(* Logix 5000 project; controller PLC_MCC1201_220AP1 vendor 1 type 14 code 164 rev 35.11; software revision 35.00; part 18 of 25 *)
(* tags used below, declared in another part *)
   B152 : DINT[50];
   B153 : DINT[20];
   B154 : DINT[20];
   B3 : DINT[102];
   C1_ACTIVE_LAMP : ALIAS FOR N54[260].0;
   C1_NTH_IN_LMP : ALIAS FOR N54[260].10;
   C1_NTH_IN_PE : ALIAS FOR N54[260].6;
   C1_NTH_IN_SS : ALIAS FOR N54[260].2;
   C1_NTH_OUT_LMP : ALIAS FOR N54[260].9;
   C1_NTH_OUT_PE : ALIAS FOR N54[260].5;
   C1_NTH_OUT_SS : ALIAS FOR N54[260].1;
   C1_STH_IN_LMP : ALIAS FOR N54[260].12;
   C1_STH_IN_PE : ALIAS FOR N54[260].8;
   C1_STH_IN_SS : ALIAS FOR N54[260].4;
   C1_STH_OUT_LMP : ALIAS FOR N54[260].11;
   C1_STH_OUT_PE : ALIAS FOR N54[260].7;
   C1_STH_OUT_SS : ALIAS FOR N54[260].3;
   C2_ACTIVE_LAMP : ALIAS FOR N54[261].0;
   C2_NTH_IN_LMP : ALIAS FOR N54[261].10;
   C2_NTH_IN_PE : ALIAS FOR N54[261].6;
   C2_NTH_IN_SS : ALIAS FOR N54[261].2;
   C2_NTH_OUT_LMP : ALIAS FOR N54[261].9;
   C2_NTH_OUT_PE : ALIAS FOR N54[261].5;
   C2_NTH_OUT_SS : ALIAS FOR N54[261].1;
   C2_STH_IN_LMP : ALIAS FOR N54[261].12;
   C2_STH_IN_PE : ALIAS FOR N54[261].8;
   C2_STH_IN_SS : ALIAS FOR N54[261].4;
   C2_STH_OUT_LMP : ALIAS FOR N54[261].11;
   C2_STH_OUT_PE : ALIAS FOR N54[261].7;
   C2_STH_OUT_SS : ALIAS FOR N54[261].3;
   C3_ACTIVE_LAMP : ALIAS FOR N54[262].0;
   C3_NTH_IN_LMP : ALIAS FOR N54[262].10;
   C3_NTH_IN_PE : ALIAS FOR N54[262].6;
   C3_NTH_IN_SS : ALIAS FOR N54[262].2;
   C3_NTH_OUT_LMP : ALIAS FOR N54[262].9;
   C3_NTH_OUT_PE : ALIAS FOR N54[262].5;
   C3_NTH_OUT_SS : ALIAS FOR N54[262].1;
   C3_STH_IN_LMP : ALIAS FOR N54[262].12;
   C3_STH_IN_PE : ALIAS FOR N54[262].8;
   C3_STH_IN_SS : ALIAS FOR N54[262].4;
   C3_STH_OUT_LMP : ALIAS FOR N54[262].11;
   C3_STH_OUT_PE : ALIAS FOR N54[262].7;
   C3_STH_OUT_SS : ALIAS FOR N54[262].3;
   C3_STP : ALIAS FOR O[35].10;
   C5 : COUNTER[100];
   C5_ACTIVE_LAMP : ALIAS FOR N54[264].0;
   C5_NTH_IN_SS : ALIAS FOR N54[264].2;
   C5_NTH_OUT_SS : ALIAS FOR N54[264].1;
   C5_STH_IN_SS : ALIAS FOR N54[264].4;
   C5_STH_OUT_SS : ALIAS FOR N54[264].3;
   CAWSV_ON_BIT_TO_WPLC : ALIAS FOR N251[900].0;
   I : INT[128];
   MADSEN_2IN_PULS : ALIAS FOR I[12].15;
   N163 : DINT[5];
   N53 : DINT[10];
   N54 : DINT[501];
   O : INT[128];
   REL_2IN_PULSE : ALIAS FOR N54[301].1;
   REL_DATA_REQ : ALIAS FOR N54[301].0;
   RELDR_ESTOP : ALIAS FOR I[80].0;
   S : INT[128];
   Status : INT;   // INT tag to retrieve Status value through GSV created during conversion
   T160 : TIMER[100];
   T4 : TIMER[100];
   T51 : TIMER[13];
   T57 : TIMER[100];
   TONY : ALIAS FOR B3[10].15;
   WASH_AK1_CON : ALIAS FOR N54[203].4;
   WASH_AK1_CR : ALIAS FOR N54[207].4;
   WASH_AK1_RET : ALIAS FOR N54[203].3;
   WASH_AK1_SV : ALIAS FOR O[36].2;
   WASH_AK1LO_CVG : ALIAS FOR N54[206].4;
   WASH_AK1UP_CVG : ALIAS FOR N54[205].4;
   WASH_AK2_CON : ALIAS FOR N54[203].6;
   WASH_AK2_CR : ALIAS FOR N54[207].5;
   WASH_AK2_RET : ALIAS FOR N54[203].5;
   WASH_AK2_SV : ALIAS FOR O[36].0;
   WASH_AK2LO_CVG : ALIAS FOR N54[206].5;
   WASH_AK2UP_CVG : ALIAS FOR N54[205].5;
   WASH_ARK_AUTO : ALIAS FOR N54[203].1;
   WASH_ARK_MANUAL : ALIAS FOR N54[203].2;
   WASH_CR_ACK : ALIAS FOR N54[207].0;
   WASH_SPY_AUTO : ALIAS FOR N54[204].1;
   WASH_SPY_MANLMP : ALIAS FOR N54[204].9;
   WASH_SPY_MANUAL : ALIAS FOR N54[204].2;
   WASH_SPY_OFF : ALIAS FOR N54[204].4;
   WASH_SPY_ON : ALIAS FOR N54[204].3;
   WATER2_ON : ALIAS FOR O[47].8;
   WATER3_CR : ALIAS FOR N54[207].6;
   WATER3_ON : ALIAS FOR O[47].9;
(* MainProgram, continued *)

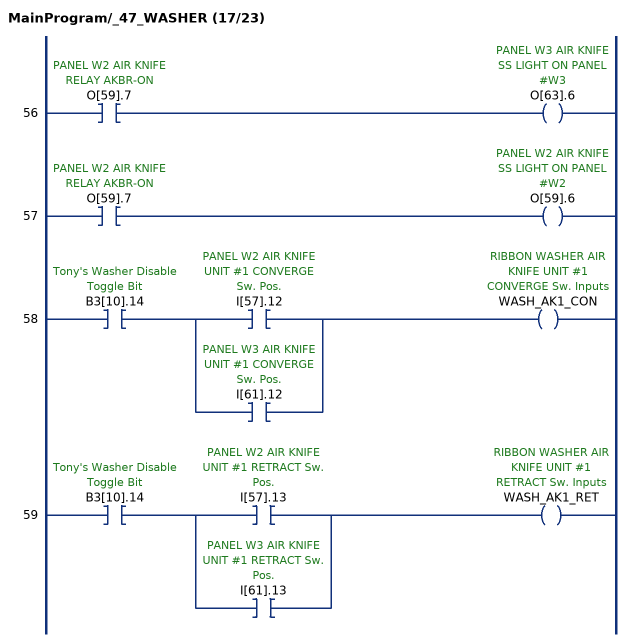
   [picture p282: MainProgram/_47_WASHER rungs 56-59]
   56: XIC(O[59].7)OTE(O[63].6);
   57: XIC(O[59].7)OTE(O[59].6);
   58: XIC(B3[10].14)[XIC(I[57].12) ,XIC(I[61].12) ]OTE(WASH_AK1_CON);
   59: XIC(B3[10].14)[XIC(I[57].13) ,XIC(I[61].13) ]OTE(WASH_AK1_RET);
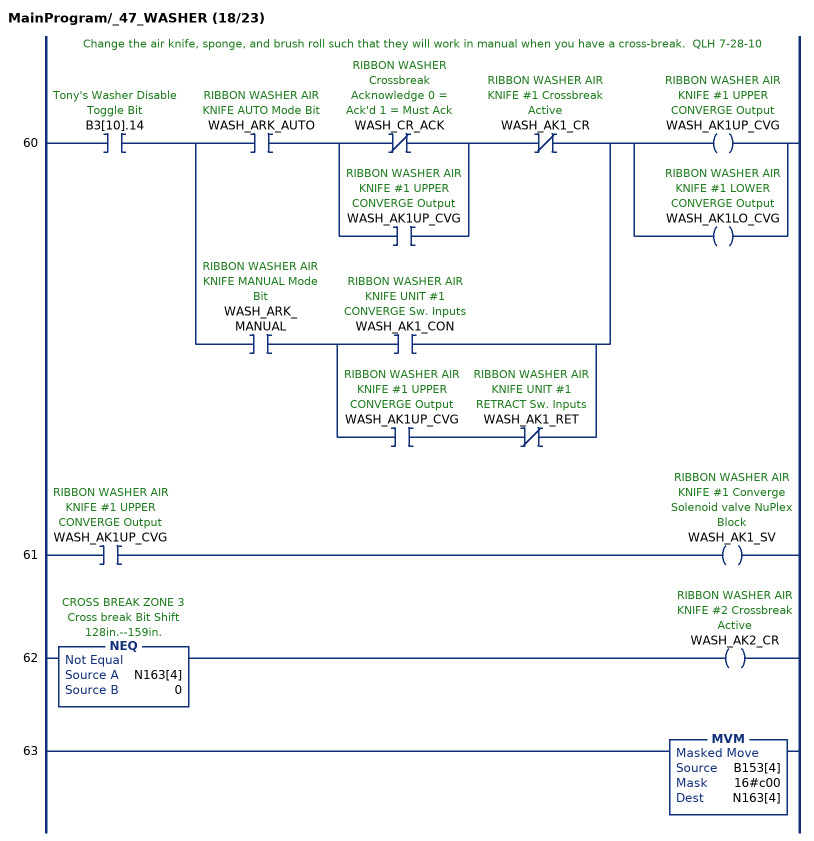
   // Change the air knife, sponge, and brush roll such that they will work in manual when you have a cross-break.  QLH 7-28-10
   60: XIC(B3[10].14)[XIC(WASH_ARK_AUTO) [XIO(WASH_CR_ACK) ,XIC(WASH_AK1UP_CVG) ] XIO(WASH_AK1_CR) ,XIC(WASH_ARK_MANUAL) [XIC(WASH_AK1_CON) ,XIC(WASH_AK1UP_CVG) XIO(WASH_AK1_RET) ] ][OTE(WASH_AK1UP_CVG) ,OTE(WASH_AK1LO_CVG) ];
   61: XIC(WASH_AK1UP_CVG)OTE(WASH_AK1_SV);
   62: NEQ(N163[4],0)OTE(WASH_AK2_CR);
   63: MVM(B153[4],16#c00,N163[4]);
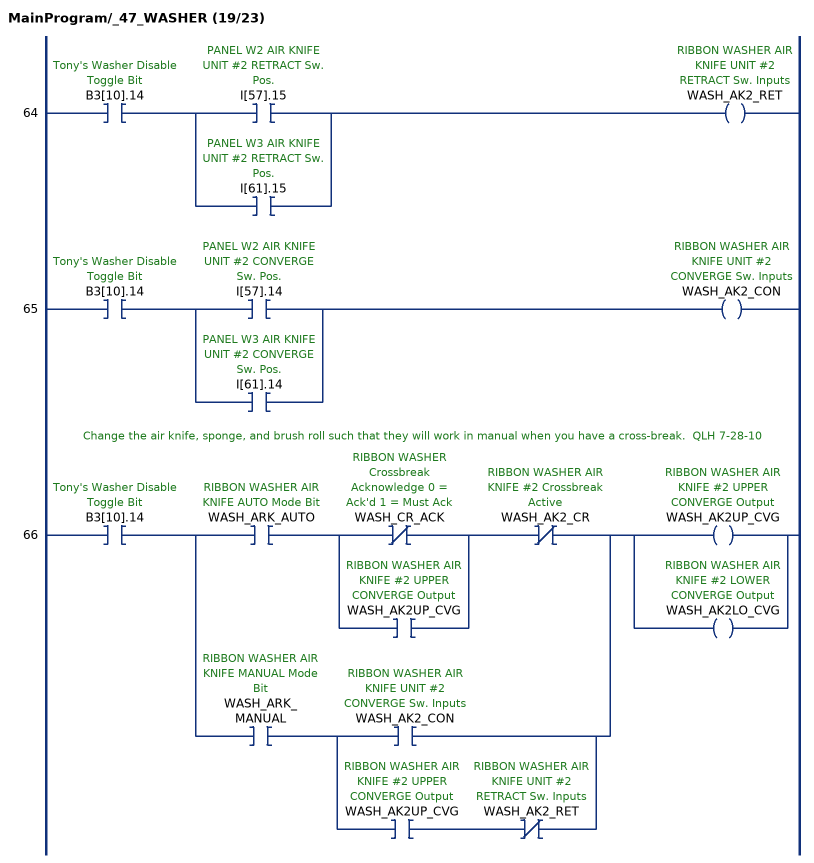
   64: XIC(B3[10].14)[XIC(I[57].15) ,XIC(I[61].15) ]OTE(WASH_AK2_RET);
   65: XIC(B3[10].14)[XIC(I[57].14) ,XIC(I[61].14) ]OTE(WASH_AK2_CON);
   // Change the air knife, sponge, and brush roll such that they will work in manual when you have a cross-break.  QLH 7-28-10
   66: XIC(B3[10].14)[XIC(WASH_ARK_AUTO) [XIO(WASH_CR_ACK) ,XIC(WASH_AK2UP_CVG) ] XIO(WASH_AK2_CR) ,XIC(WASH_ARK_MANUAL) [XIC(WASH_AK2_CON) ,XIC(WASH_AK2UP_CVG) XIO(WASH_AK2_RET) ] ][OTE(WASH_AK2UP_CVG) ,OTE(WASH_AK2LO_CVG) ];
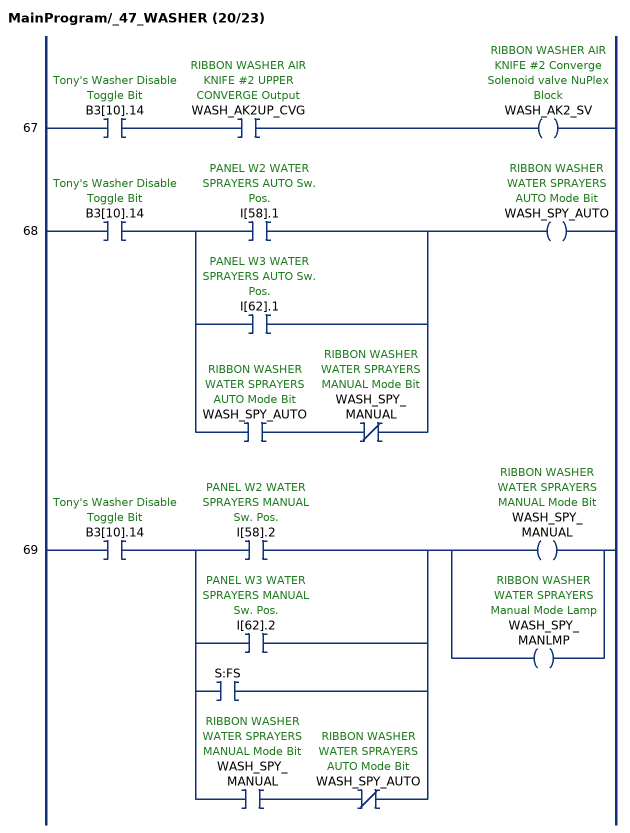
   67: XIC(B3[10].14)XIC(WASH_AK2UP_CVG)OTE(WASH_AK2_SV);
   68: XIC(B3[10].14)[[XIC(I[58].1) ,XIC(I[62].1) ] ,XIC(WASH_SPY_AUTO) XIO(WASH_SPY_MANUAL) ]OTE(WASH_SPY_AUTO);
   69: XIC(B3[10].14)[[XIC(I[58].2) ,XIC(I[62].2) ,XIC(S:FS) ] ,XIC(WASH_SPY_MANUAL) XIO(WASH_SPY_AUTO) ][OTE(WASH_SPY_MANUAL) ,OTE(WASH_SPY_MANLMP) ];
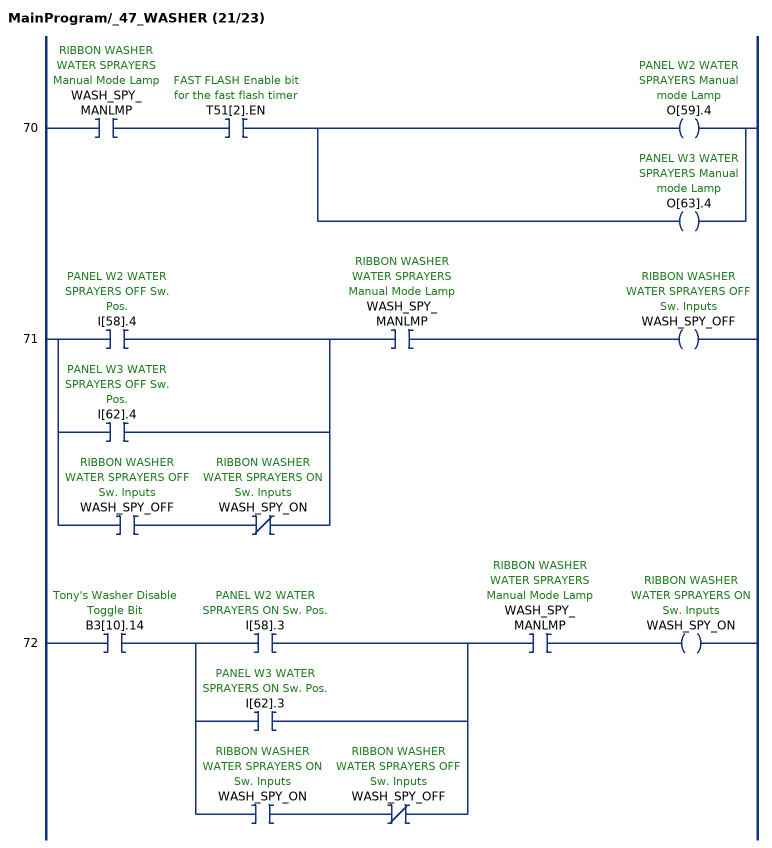
   70: XIC(WASH_SPY_MANLMP)XIC(T51[2].EN)[OTE(O[59].4) ,OTE(O[63].4) ];
   71: [[XIC(I[58].4) ,XIC(I[62].4) ] ,XIC(WASH_SPY_OFF) XIO(WASH_SPY_ON) ]XIC(WASH_SPY_MANLMP)OTE(WASH_SPY_OFF);
   72: XIC(B3[10].14)[[XIC(I[58].3) ,XIC(I[62].3) ] ,XIC(WASH_SPY_ON) XIO(WASH_SPY_OFF) ]XIC(WASH_SPY_MANLMP)OTE(WASH_SPY_ON);
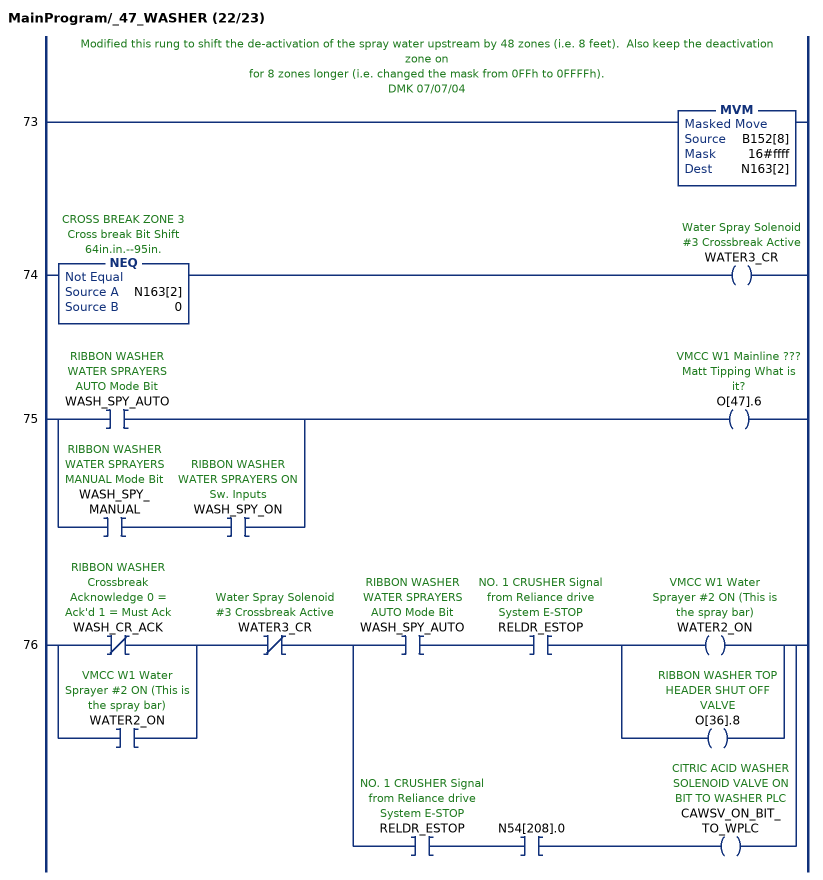
   // Modified this rung to shift the de-activation of the spray water upstream by 48 zones (i.e. 8 feet).  Also keep the deactivation zone on
   // for 8 zones longer (i.e. changed the mask from 0FFh to 0FFFFh).
   // DMK 07/07/04
   73: MVM(B152[8],16#ffff,N163[2]);
   74: NEQ(N163[2],0)OTE(WATER3_CR);
   75: [XIC(WASH_SPY_AUTO) ,XIC(WASH_SPY_MANUAL) XIC(WASH_SPY_ON) ]OTE(O[47].6);
   76: [XIO(WASH_CR_ACK) ,XIC(WATER2_ON) ]XIO(WATER3_CR)[XIC(WASH_SPY_AUTO) XIC(RELDR_ESTOP) [OTE(WATER2_ON) ,OTE(O[36].8) ] ,XIC(RELDR_ESTOP) XIC(N54[208].0) OTE(CAWSV_ON_BIT_TO_WPLC) ];
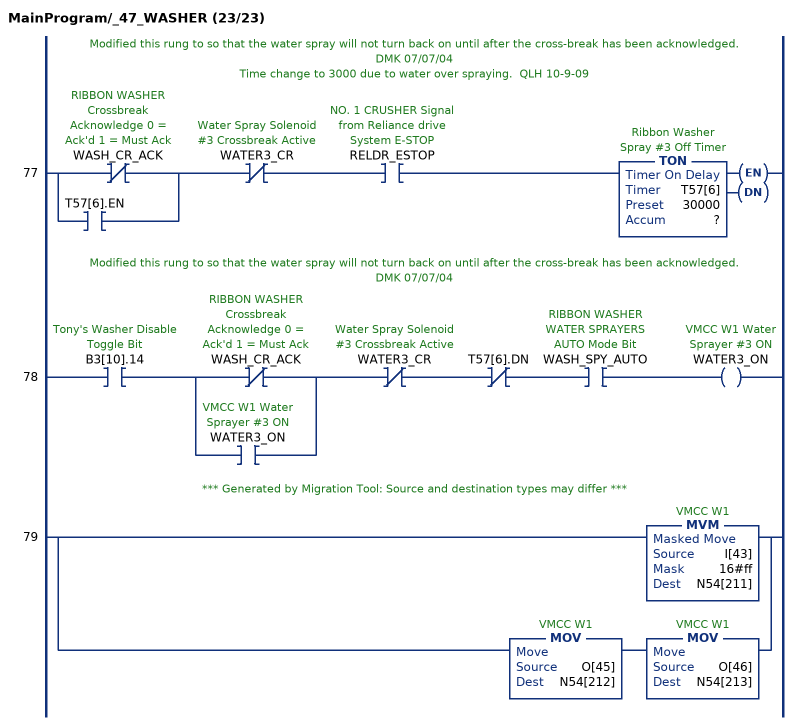
   // Modified this rung to so that the water spray will not turn back on until after the cross-break has been acknowledged.
   // DMK 07/07/04
   // Time change to 3000 due to water over spraying.  QLH 10-9-09
   77: [XIO(WASH_CR_ACK) ,XIC(T57[6].EN) ]XIO(WATER3_CR)XIC(RELDR_ESTOP)TON(T57[6],?,?);
   // Modified this rung to so that the water spray will not turn back on until after the cross-break has been acknowledged.
   // DMK 07/07/04
   78: XIC(B3[10].14)[XIO(WASH_CR_ACK) ,XIC(WATER3_ON) ]XIO(WATER3_CR)XIO(T57[6].DN)XIC(WASH_SPY_AUTO)OTE(WATER3_ON);
   // *** Generated by Migration Tool: Source and destination types may differ ***
   79: [MVM(I[43],16#ff,N54[211]) ,MOV(O[45],N54[212]) MOV(O[46],N54[213]) ];
END_ROUTINE

ROUTINE _48_IMAGE   (* ladder *)
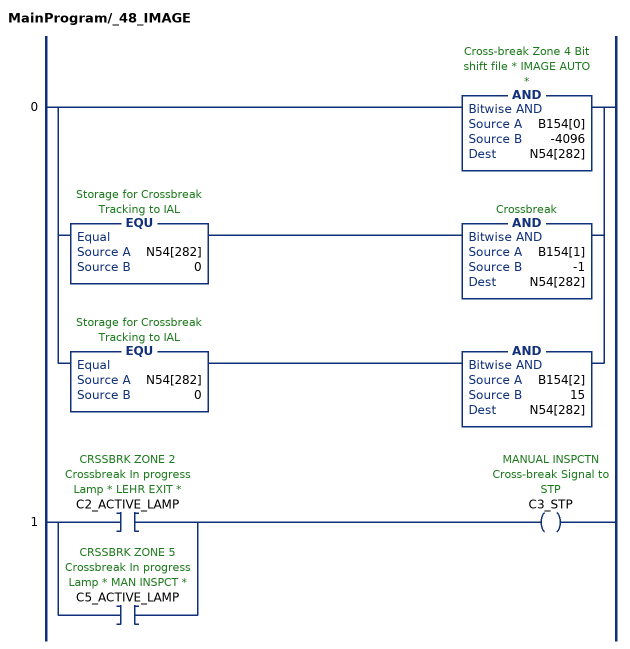
   0: [AND(B154[0],-4096,N54[282]) ,EQU(N54[282],0) AND(B154[1],-1,N54[282]) ,EQU(N54[282],0) AND(B154[2],15,N54[282]) ];
   1: [XIC(C2_ACTIVE_LAMP) ,XIC(C5_ACTIVE_LAMP) ]OTE(C3_STP);
END_ROUTINE

ROUTINE _49_INSP_REL   (* ladder *)
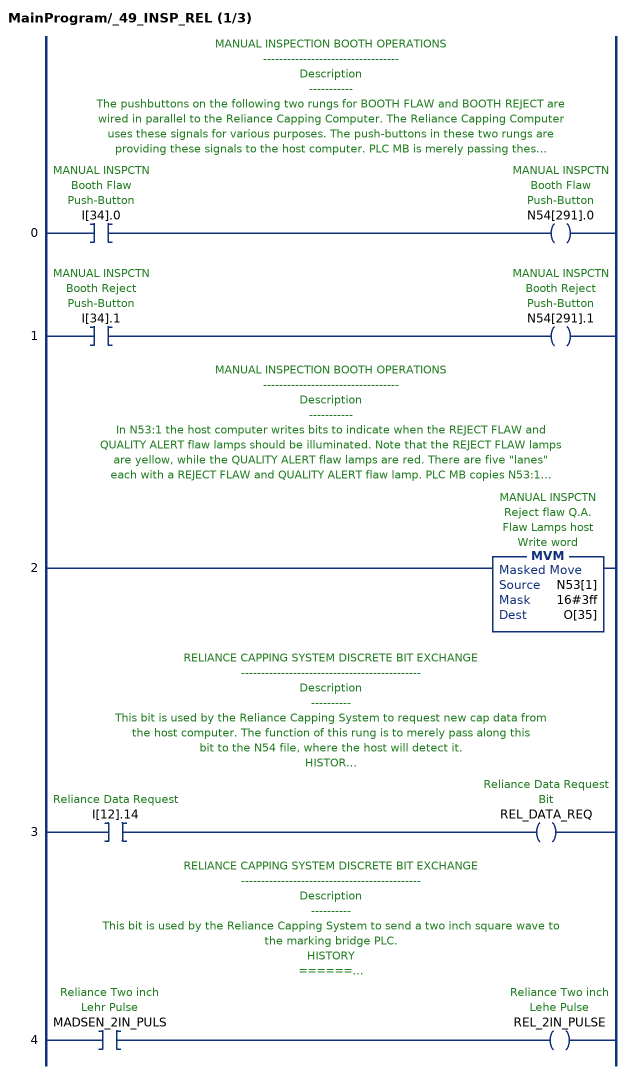
   // MANUAL INSPECTION BOOTH OPERATIONS
   // ----------------------------------
   // Description
   // -----------
   // The pushbuttons on the following two rungs for BOOTH FLAW and BOOTH REJECT are
   // wired in parallel to the Reliance Capping Computer. The Reliance Capping Computer
   // uses these signals for various purposes. The push-buttons in these two rungs are
   // providing these signals to the host computer. PLC MB is merely passing these
   // signals along to the host computer.
   // HISTORY
   // =======
   // Date       Description                                                Programmer
   // ----       -----------                                                ----------
   // 3/11/96    Added this rung and comments.                                WAS
   0: XIC(I[34].0)OTE(N54[291].0);
   1: XIC(I[34].1)OTE(N54[291].1);
   // MANUAL INSPECTION BOOTH OPERATIONS
   // ----------------------------------
   // Description
   // -----------
   // In N53:1 the host computer writes bits to indicate when the REJECT FLAW and
   // QUALITY ALERT flaw lamps should be illuminated. Note that the REJECT FLAW lamps
   // are yellow, while the QUALITY ALERT flaw lamps are red. There are five "lanes"
   // each with a REJECT FLAW and QUALITY ALERT flaw lamp. PLC MB copies N53:1,
   // the host write area, to O:043, the actual output word for the lamps.
   // HISTORY
   // =======
   // Date       Description                                                Programmer
   // ----       -----------                                                ----------
   // 3/11/96    Added this rung and comments.                                WAS
   2: MVM(N53[1],16#3ff,O[35]);
   // RELIANCE CAPPING SYSTEM DISCRETE BIT EXCHANGE
   // ---------------------------------------------
   // Description
   // ----------
   // This bit is used by the Reliance Capping System to request new cap data from
   // the host computer. The function of this rung is to merely pass along this
   // bit to the N54 file, where the host will detect it.
   // HISTORY
   // =======
   // Date       Description                                                Programmer
   // ----       -----------                                                ----------
   // 3/11/96    Discussed issue with Steve Sutter. Elected to locate This    WAS
   //            bit in local rack in case timing becomes critical.
   // 3/11/96    Added this rung and comments.                                WAS
   3: XIC(I[12].14)OTE(REL_DATA_REQ);
   // RELIANCE CAPPING SYSTEM DISCRETE BIT EXCHANGE
   // ---------------------------------------------
   // Description
   // ----------
   // This bit is used by the Reliance Capping System to send a two inch square wave to
   // the marking bridge PLC.
   // HISTORY
   // =======
   // Date       Description                                                Programmer
   // ----       -----------                                                ----------
   // 3/11/96    Discussed issue with Steve Sutter. Elected to locate This    WAS
   //            bit in local rack in case timing becomes critical.
   // 3/11/96    Added this rung and comments.                                WAS
   4: XIC(MADSEN_2IN_PULS)OTE(REL_2IN_PULSE);
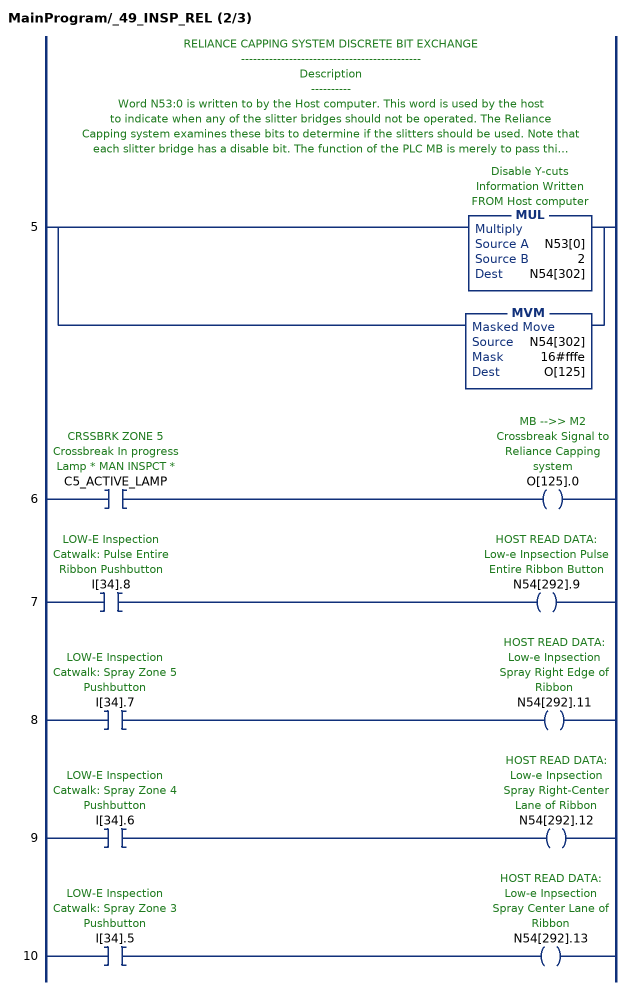
   // RELIANCE CAPPING SYSTEM DISCRETE BIT EXCHANGE
   // ---------------------------------------------
   // Description
   // ----------
   // Word N53:0 is written to by the Host computer. This word is used by the host
   // to indicate when any of the slitter bridges should not be operated. The Reliance
   // Capping system examines these bits to determine if the slitters should be used. Note that
   // each slitter bridge has a disable bit. The function of the PLC MB is merely to pass this
   // data along from the Host computer to the Reliance Capping System.
   // HISTORY
   // =======
   // Date       Description                                                Programmer
   // ----       -----------                                                ----------
   // 3/11/96    Added this rung and comments.                                WAS
   5: [MUL(N53[0],2,N54[302]) ,MVM(N54[302],16#fffe,O[125]) ];
   6: XIC(C5_ACTIVE_LAMP)OTE(O[125].0);
   7: XIC(I[34].8)OTE(N54[292].9);
   8: XIC(I[34].7)OTE(N54[292].11);
   9: XIC(I[34].6)OTE(N54[292].12);
   10: XIC(I[34].5)OTE(N54[292].13);
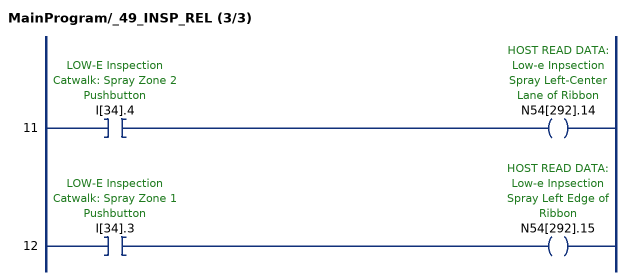
   11: XIC(I[34].4)OTE(N54[292].14);
   12: XIC(I[34].3)OTE(N54[292].15);
END_ROUTINE

ROUTINE _50_I_O_REMAP   (* ladder *)
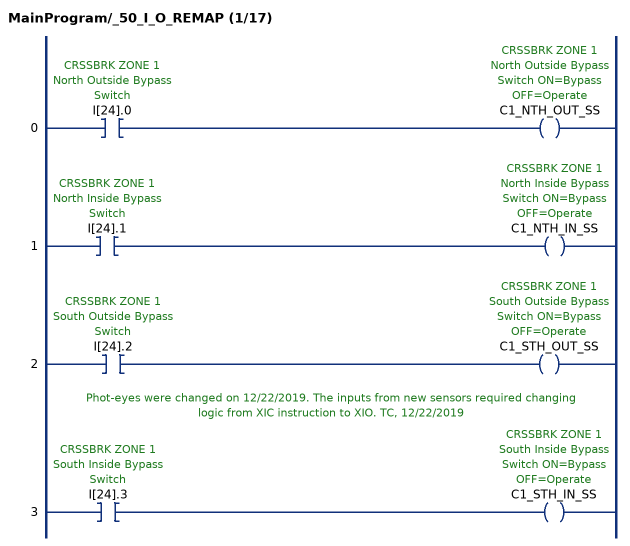
   0: XIC(I[24].0)OTE(C1_NTH_OUT_SS);
   1: XIC(I[24].1)OTE(C1_NTH_IN_SS);
   2: XIC(I[24].2)OTE(C1_STH_OUT_SS);
   // Phot-eyes were changed on 12/22/2019. The inputs from new sensors required changing logic from XIC instruction to XIO. TC, 12/22/2019
   3: XIC(I[24].3)OTE(C1_STH_IN_SS);
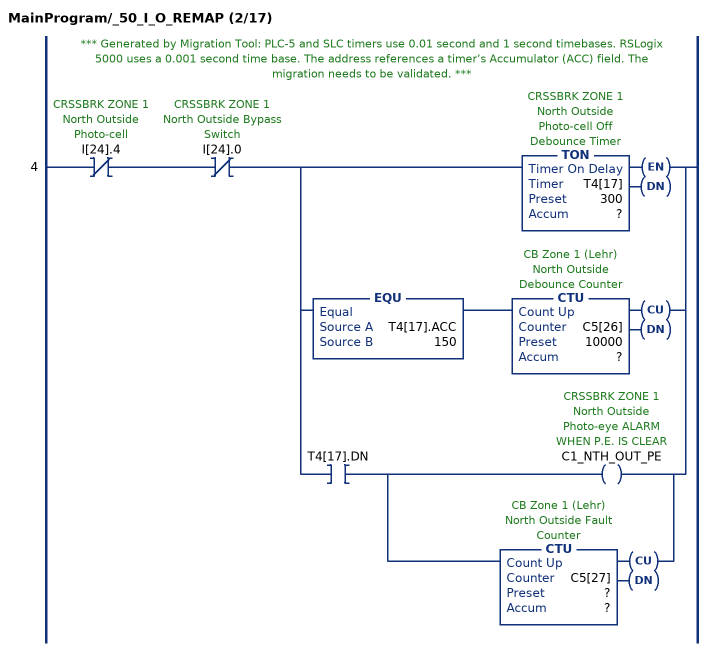
   // *** Generated by Migration Tool: PLC-5 and SLC timers use 0.01 second and 1 second timebases. RSLogix 5000 uses a 0.001 second time base. The address references a timer’s Accumulator (ACC) field. The migration needs to be validated. ***
   4: XIO(I[24].4)XIO(I[24].0)[TON(T4[17],?,?) ,EQU(T4[17].ACC,150) CTU(C5[26],?,?) ,XIC(T4[17].DN) [OTE(C1_NTH_OUT_PE) ,CTU(C5[27],?,?) ] ];
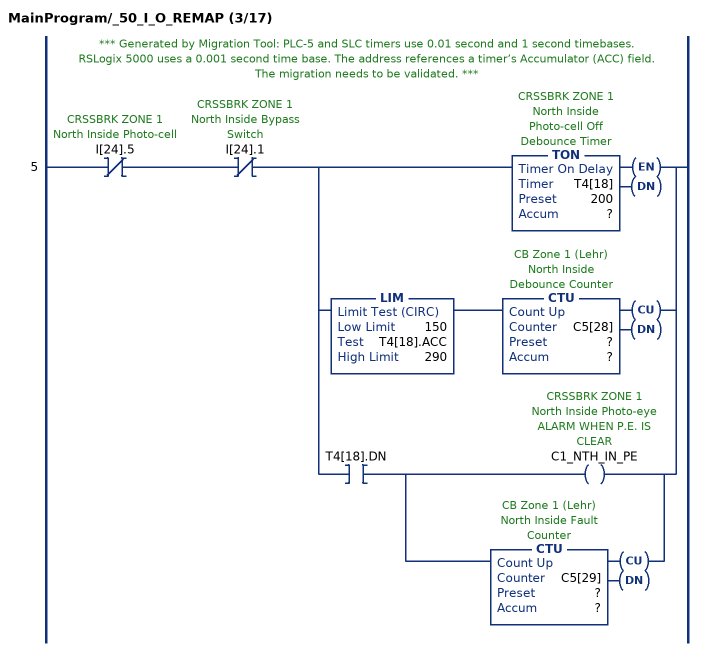
   // *** Generated by Migration Tool: PLC-5 and SLC timers use 0.01 second and 1 second timebases. RSLogix 5000 uses a 0.001 second time base. The address references a timer’s Accumulator (ACC) field. The migration needs to be validated. ***
   5: XIO(I[24].5)XIO(I[24].1)[TON(T4[18],?,?) ,LIM(150,T4[18].ACC,290) CTU(C5[28],?,?) ,XIC(T4[18].DN) [OTE(C1_NTH_IN_PE) ,CTU(C5[29],?,?) ] ];
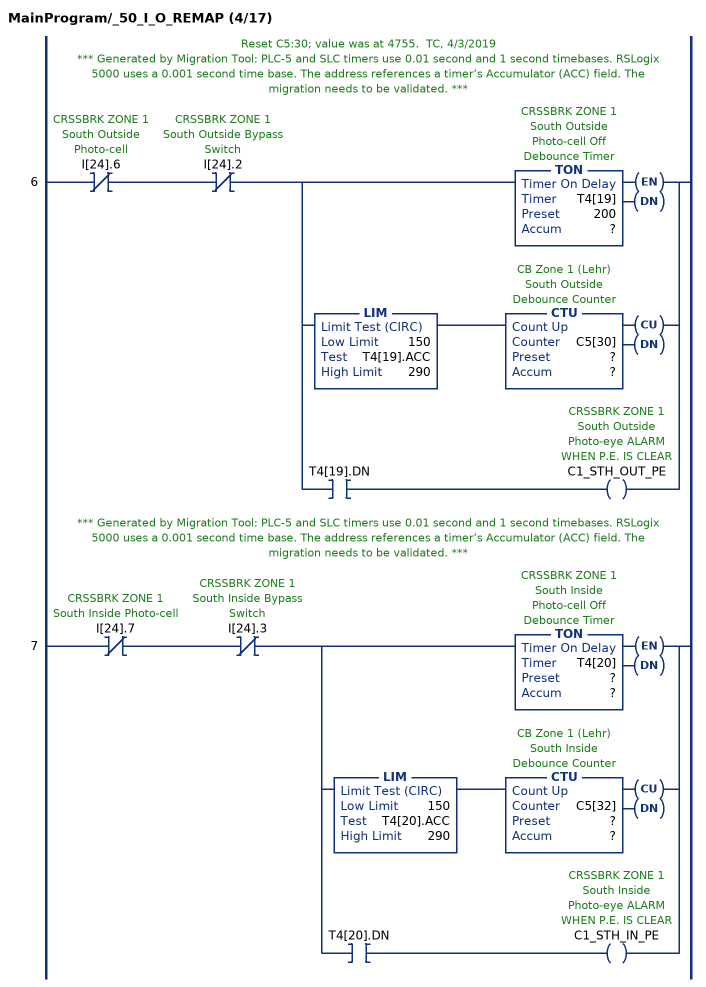
   // Reset C5:30; value was at 4755.  TC, 4/3/2019
   // *** Generated by Migration Tool: PLC-5 and SLC timers use 0.01 second and 1 second timebases. RSLogix 5000 uses a 0.001 second time base. The address references a timer’s Accumulator (ACC) field. The migration needs to be validated. ***
   6: XIO(I[24].6)XIO(I[24].2)[TON(T4[19],?,?) ,LIM(150,T4[19].ACC,290) CTU(C5[30],?,?) ,XIC(T4[19].DN) OTE(C1_STH_OUT_PE) ];
   // *** Generated by Migration Tool: PLC-5 and SLC timers use 0.01 second and 1 second timebases. RSLogix 5000 uses a 0.001 second time base. The address references a timer’s Accumulator (ACC) field. The migration needs to be validated. ***
   7: XIO(I[24].7)XIO(I[24].3)[TON(T4[20],?,?) ,LIM(150,T4[20].ACC,290) CTU(C5[32],?,?) ,XIC(T4[20].DN) OTE(C1_STH_IN_PE) ];
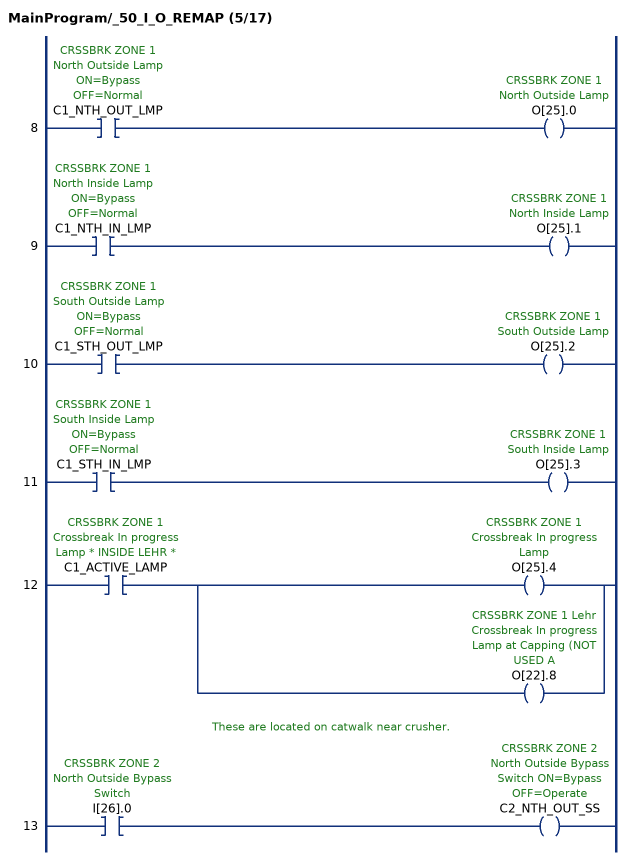
   8: XIC(C1_NTH_OUT_LMP)OTE(O[25].0);
   9: XIC(C1_NTH_IN_LMP)OTE(O[25].1);
   10: XIC(C1_STH_OUT_LMP)OTE(O[25].2);
   11: XIC(C1_STH_IN_LMP)OTE(O[25].3);
   12: XIC(C1_ACTIVE_LAMP)[OTE(O[25].4) ,OTE(O[22].8) ];
   // These are located on catwalk near crusher.
   13: XIC(I[26].0)OTE(C2_NTH_OUT_SS);
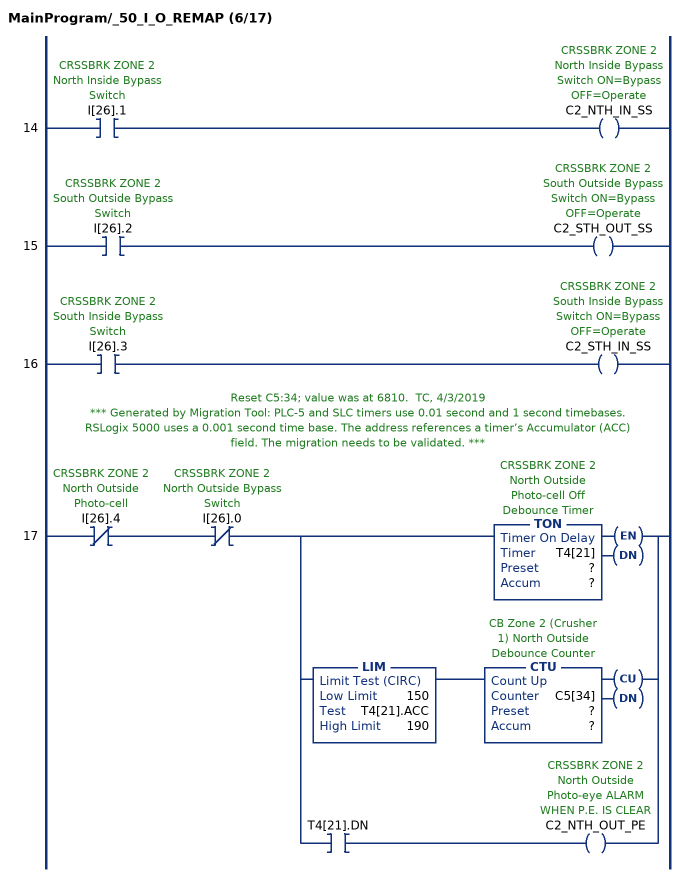
   14: XIC(I[26].1)OTE(C2_NTH_IN_SS);
   15: XIC(I[26].2)OTE(C2_STH_OUT_SS);
   16: XIC(I[26].3)OTE(C2_STH_IN_SS);
   // Reset C5:34; value was at 6810.  TC, 4/3/2019
   // *** Generated by Migration Tool: PLC-5 and SLC timers use 0.01 second and 1 second timebases. RSLogix 5000 uses a 0.001 second time base. The address references a timer’s Accumulator (ACC) field. The migration needs to be validated. ***
   17: XIO(I[26].4)XIO(I[26].0)[TON(T4[21],?,?) ,LIM(150,T4[21].ACC,190) CTU(C5[34],?,?) ,XIC(T4[21].DN) OTE(C2_NTH_OUT_PE) ];
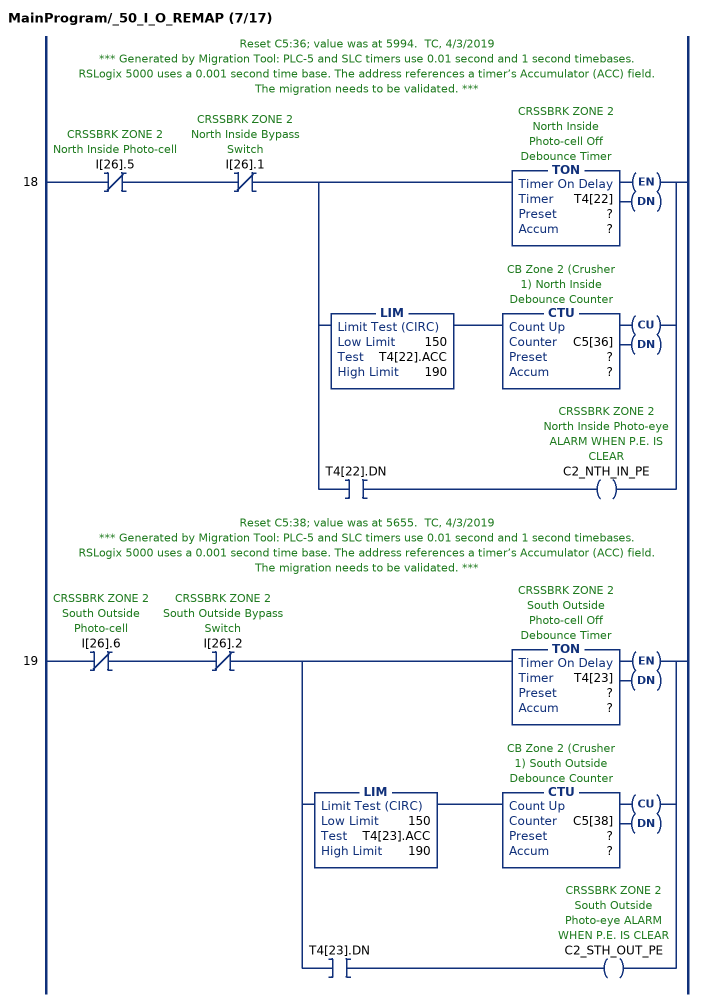
   // Reset C5:36; value was at 5994.  TC, 4/3/2019
   // *** Generated by Migration Tool: PLC-5 and SLC timers use 0.01 second and 1 second timebases. RSLogix 5000 uses a 0.001 second time base. The address references a timer’s Accumulator (ACC) field. The migration needs to be validated. ***
   18: XIO(I[26].5)XIO(I[26].1)[TON(T4[22],?,?) ,LIM(150,T4[22].ACC,190) CTU(C5[36],?,?) ,XIC(T4[22].DN) OTE(C2_NTH_IN_PE) ];
   // Reset C5:38; value was at 5655.  TC, 4/3/2019
   // *** Generated by Migration Tool: PLC-5 and SLC timers use 0.01 second and 1 second timebases. RSLogix 5000 uses a 0.001 second time base. The address references a timer’s Accumulator (ACC) field. The migration needs to be validated. ***
   19: XIO(I[26].6)XIO(I[26].2)[TON(T4[23],?,?) ,LIM(150,T4[23].ACC,190) CTU(C5[38],?,?) ,XIC(T4[23].DN) OTE(C2_STH_OUT_PE) ];
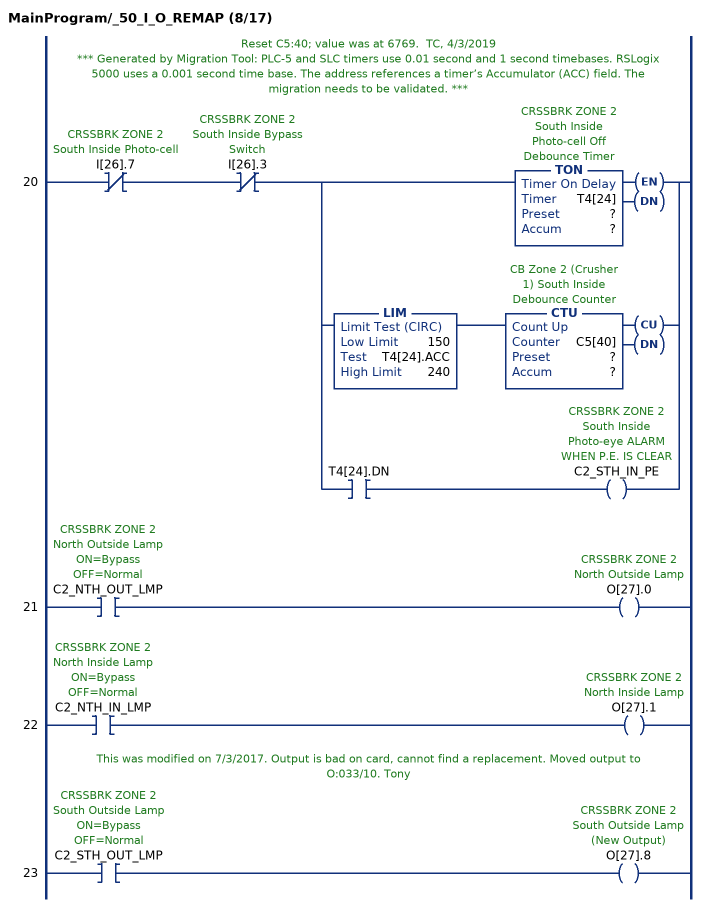
   // Reset C5:40; value was at 6769.  TC, 4/3/2019
   // *** Generated by Migration Tool: PLC-5 and SLC timers use 0.01 second and 1 second timebases. RSLogix 5000 uses a 0.001 second time base. The address references a timer’s Accumulator (ACC) field. The migration needs to be validated. ***
   20: XIO(I[26].7)XIO(I[26].3)[TON(T4[24],?,?) ,LIM(150,T4[24].ACC,240) CTU(C5[40],?,?) ,XIC(T4[24].DN) OTE(C2_STH_IN_PE) ];
   21: XIC(C2_NTH_OUT_LMP)OTE(O[27].0);
   22: XIC(C2_NTH_IN_LMP)OTE(O[27].1);
   // This was modified on 7/3/2017. Output is bad on card, cannot find a replacement. Moved output to O:033/10. Tony
   23: XIC(C2_STH_OUT_LMP)OTE(O[27].8);
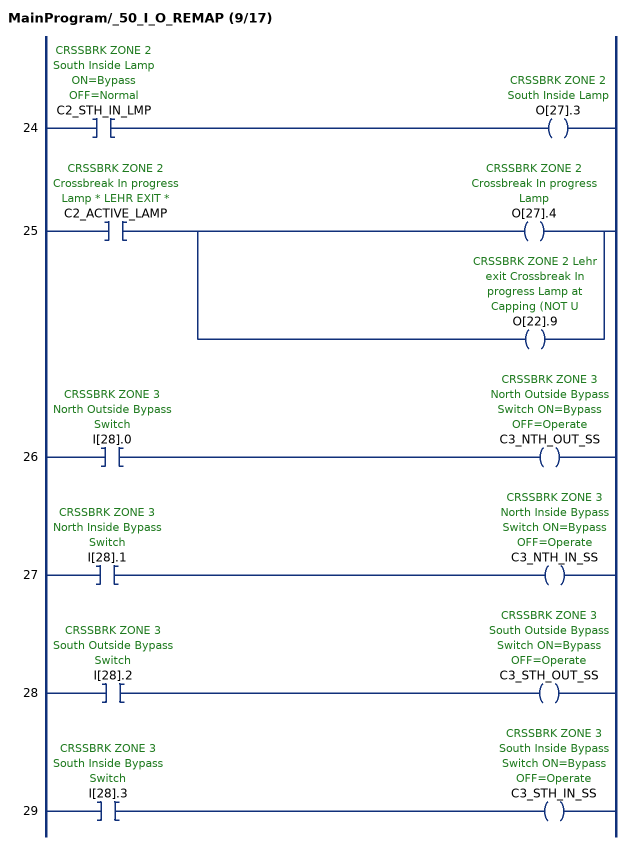
   24: XIC(C2_STH_IN_LMP)OTE(O[27].3);
   25: XIC(C2_ACTIVE_LAMP)[OTE(O[27].4) ,OTE(O[22].9) ];
   26: XIC(I[28].0)OTE(C3_NTH_OUT_SS);
   27: XIC(I[28].1)OTE(C3_NTH_IN_SS);
   28: XIC(I[28].2)OTE(C3_STH_OUT_SS);
   29: XIC(I[28].3)OTE(C3_STH_IN_SS);
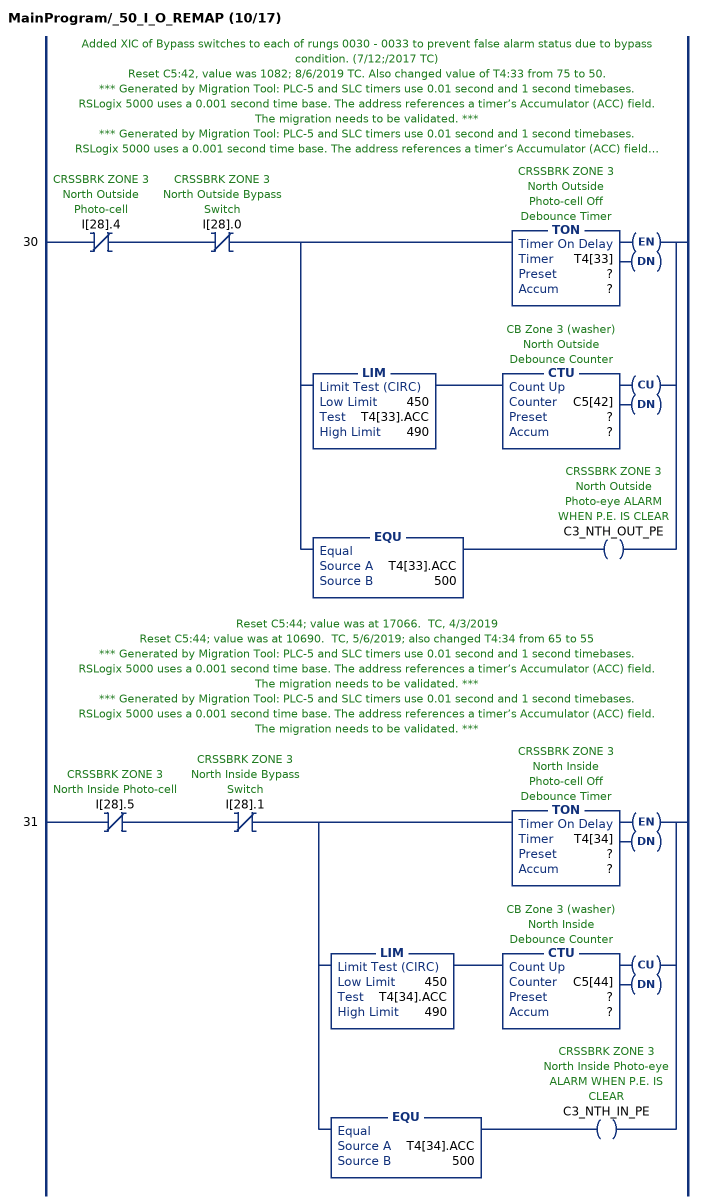
   // Added XIC of Bypass switches to each of rungs 0030 - 0033 to prevent false alarm status due to bypass condition. (7/12;/2017 TC)
   //                                                                                                                                                                    Reset C5:42, value was 1082; 8/6/2019 TC. Also changed value of T4:33 from 75 to 50.
   // *** Generated by Migration Tool: PLC-5 and SLC timers use 0.01 second and 1 second timebases. RSLogix 5000 uses a 0.001 second time base. The address references a timer’s Accumulator (ACC) field. The migration needs to be validated. ***
   // *** Generated by Migration Tool: PLC-5 and SLC timers use 0.01 second and 1 second timebases. RSLogix 5000 uses a 0.001 second time base. The address references a timer’s Accumulator (ACC) field. The migration needs to be validated. ***
   30: XIO(I[28].4)XIO(I[28].0)[TON(T4[33],?,?) ,LIM(450,T4[33].ACC,490) CTU(C5[42],?,?) ,EQU(T4[33].ACC,500) OTE(C3_NTH_OUT_PE) ];
   // Reset C5:44; value was at 17066.  TC, 4/3/2019
   //                                                                                                                                                                                      Reset C5:44; value was at 10690.  TC, 5/6/2019; also changed T4:34 from 65 to 55
   // *** Generated by Migration Tool: PLC-5 and SLC timers use 0.01 second and 1 second timebases. RSLogix 5000 uses a 0.001 second time base. The address references a timer’s Accumulator (ACC) field. The migration needs to be validated. ***
   // *** Generated by Migration Tool: PLC-5 and SLC timers use 0.01 second and 1 second timebases. RSLogix 5000 uses a 0.001 second time base. The address references a timer’s Accumulator (ACC) field. The migration needs to be validated. ***
   31: XIO(I[28].5)XIO(I[28].1)[TON(T4[34],?,?) ,LIM(450,T4[34].ACC,490) CTU(C5[44],?,?) ,EQU(T4[34].ACC,500) OTE(C3_NTH_IN_PE) ];
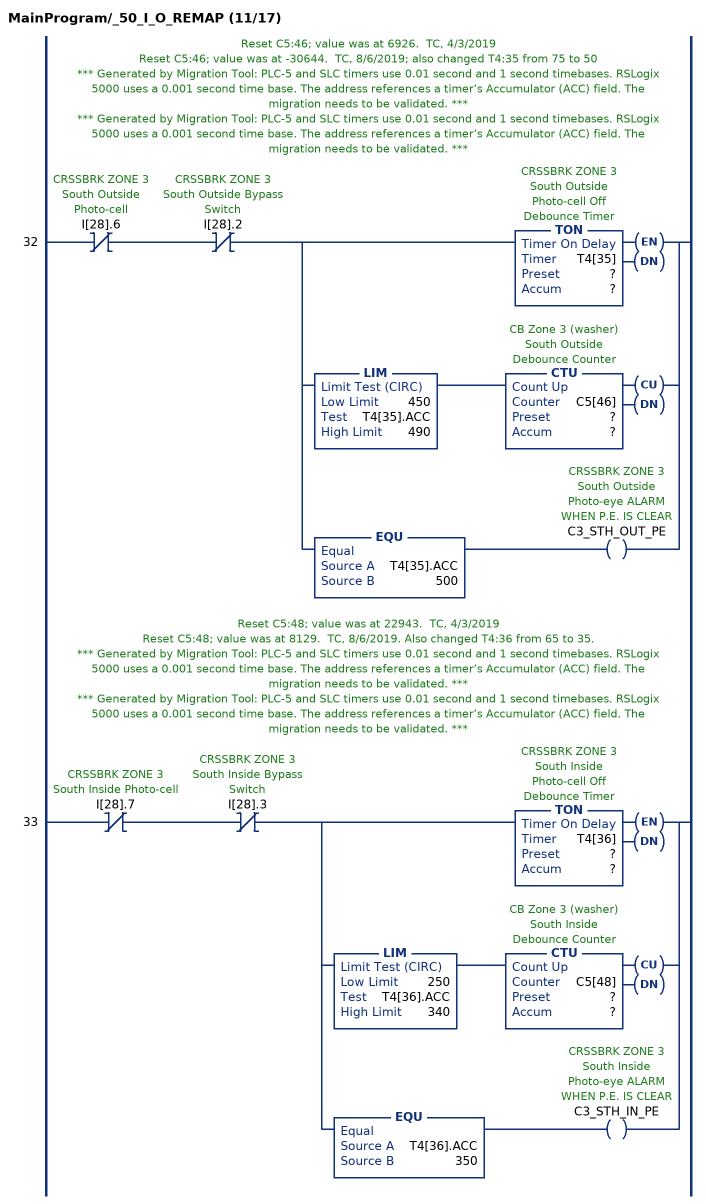
   // Reset C5:46; value was at 6926.  TC, 4/3/2019
   //                                                                                                                                                                                                  Reset C5:46; value was at -30644.  TC, 8/6/2019; also changed T4:35 from 75 to 50
   // *** Generated by Migration Tool: PLC-5 and SLC timers use 0.01 second and 1 second timebases. RSLogix 5000 uses a 0.001 second time base. The address references a timer’s Accumulator (ACC) field. The migration needs to be validated. ***
   // *** Generated by Migration Tool: PLC-5 and SLC timers use 0.01 second and 1 second timebases. RSLogix 5000 uses a 0.001 second time base. The address references a timer’s Accumulator (ACC) field. The migration needs to be validated. ***
   32: XIO(I[28].6)XIO(I[28].2)[TON(T4[35],?,?) ,LIM(450,T4[35].ACC,490) CTU(C5[46],?,?) ,EQU(T4[35].ACC,500) OTE(C3_STH_OUT_PE) ];
   // Reset C5:48; value was at 22943.  TC, 4/3/2019
   //                                                                                                                                                                      Reset C5:48; value was at 8129.  TC, 8/6/2019. Also changed T4:36 from 65 to 35.
   // *** Generated by Migration Tool: PLC-5 and SLC timers use 0.01 second and 1 second timebases. RSLogix 5000 uses a 0.001 second time base. The address references a timer’s Accumulator (ACC) field. The migration needs to be validated. ***
   // *** Generated by Migration Tool: PLC-5 and SLC timers use 0.01 second and 1 second timebases. RSLogix 5000 uses a 0.001 second time base. The address references a timer’s Accumulator (ACC) field. The migration needs to be validated. ***
   33: XIO(I[28].7)XIO(I[28].3)[TON(T4[36],?,?) ,LIM(250,T4[36].ACC,340) CTU(C5[48],?,?) ,EQU(T4[36].ACC,350) OTE(C3_STH_IN_PE) ];
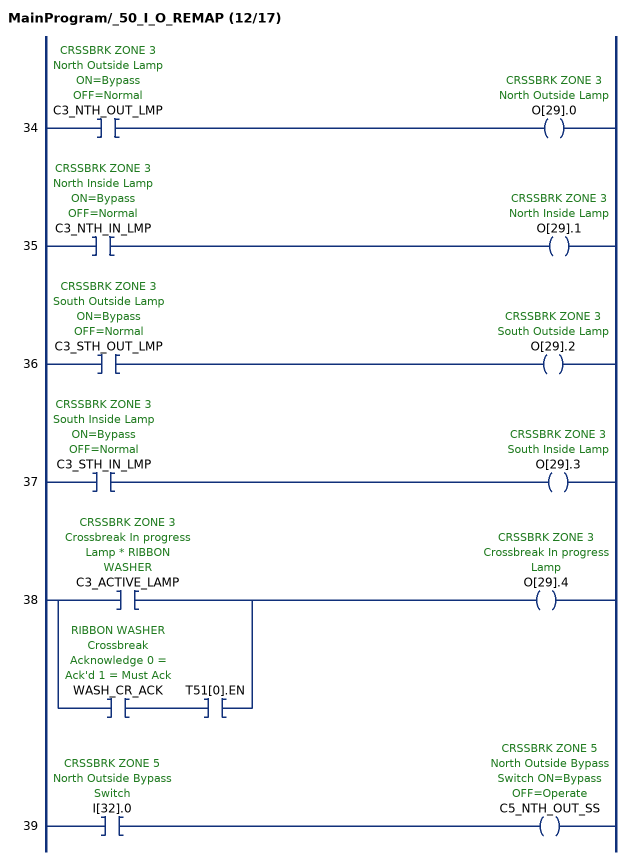
   34: XIC(C3_NTH_OUT_LMP)OTE(O[29].0);
   35: XIC(C3_NTH_IN_LMP)OTE(O[29].1);
   36: XIC(C3_STH_OUT_LMP)OTE(O[29].2);
   37: XIC(C3_STH_IN_LMP)OTE(O[29].3);
   38: [XIC(C3_ACTIVE_LAMP) ,XIC(WASH_CR_ACK) XIC(T51[0].EN) ]OTE(O[29].4);
   39: XIC(I[32].0)OTE(C5_NTH_OUT_SS);
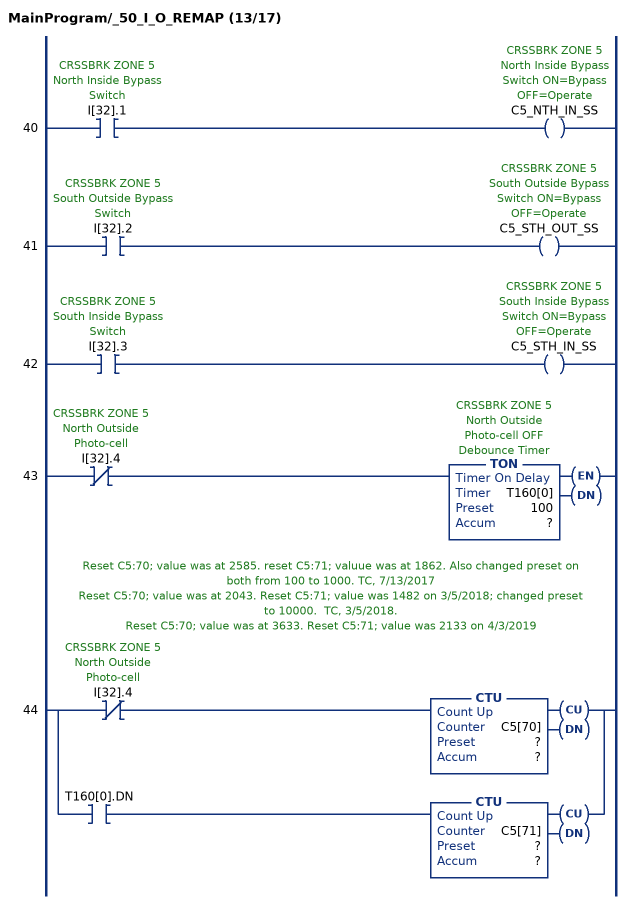
   40: XIC(I[32].1)OTE(C5_NTH_IN_SS);
   41: XIC(I[32].2)OTE(C5_STH_OUT_SS);
   42: XIC(I[32].3)OTE(C5_STH_IN_SS);
   43: XIO(I[32].4)TON(T160[0],?,?);
   // Reset C5:70; value was at 2585. reset C5:71; valuue was at 1862. Also changed preset on both from 100 to 1000. TC, 7/13/2017
   //                                                                                                                                                            Reset C5:70; value was at 2043. Reset C5:71; value was 1482 on 3/5/2018; changed preset to 10000.  TC, 3/5/2018.
   //                                                                                                                                                                              Reset C5:70; value was at 3633. Reset C5:71; value was 2133 on 4/3/2019
   44: [XIO(I[32].4) CTU(C5[70],?,?) ,XIC(T160[0].DN) CTU(C5[71],?,?) ];
